   15675: 'Mixinghead 07: Connection 02: Pressure recording: Measuring value outside measuring range', class Mixing Head Warning, trigger "Mixinghead_Pressure_MH7_Con2_DBW320" bit 8
   15676: 'Mixinghead 07: Connection 02: Pressure recording: Warning, value exceeded', class Mixing Head Warning, trigger "Mixinghead_Pressure_MH7_Con2_DBW320" bit 9
   15677: 'Mixinghead 07: Connection 02: Pressure recording: Warning, value undershot', class Mixing Head Warning, trigger "Mixinghead_Pressure_MH7_Con2_DBW320" bit 10
   15678: 'Mixinghead 07: Connection 02: Pressure recording: Fault, value exceeded', class Mixing Head Errors, trigger "Mixinghead_Pressure_MH7_Con2_DBW320" bit 11
   15679: 'Mixinghead 07: Connection 02: Pressure recording: Fault, value undershot', class Mixing Head Errors, trigger "Mixinghead_Pressure_MH7_Con2_DBW320" bit 12
   15680: 'Mixinghead 07: Connection 03: Pressure recording: Measuring value outside measuring range', class Mixing Head Warning, trigger "Mixinghead_Pressure_MH7_Con3_DBW354" bit 8
   15681: 'Mixinghead 07: Connection 03: Pressure recording: Warning, value exceeded', class Mixing Head Warning, trigger "Mixinghead_Pressure_MH7_Con3_DBW354" bit 9
   15682: 'Mixinghead 07: Connection 03: Pressure recording: Warning, value undershot', class Mixing Head Warning, trigger "Mixinghead_Pressure_MH7_Con3_DBW354" bit 10
   15683: 'Mixinghead 07: Connection 03: Pressure recording: Fault, value exceeded', class Mixing Head Errors, trigger "Mixinghead_Pressure_MH7_Con3_DBW354" bit 11
   15684: 'Mixinghead 07: Connection 03: Pressure recording: Fault, value undershot', class Mixing Head Errors, trigger "Mixinghead_Pressure_MH7_Con3_DBW354" bit 12
   15685: 'Mixinghead 07: Connection 04: Pressure recording: Measuring value outside measuring range', class Mixing Head Warning, trigger "Mixinghead_Pressure_MH7_Con4_DBW388" bit 8
   15686: 'Mixinghead 07: Connection 04: Pressure recording: Warning, value exceeded', class Mixing Head Warning, trigger "Mixinghead_Pressure_MH7_Con4_DBW388" bit 9
   15687: 'Mixinghead 07: Connection 04: Pressure recording: Warning, value undershot', class Mixing Head Warning, trigger "Mixinghead_Pressure_MH7_Con4_DBW388" bit 10
   15688: 'Mixinghead 07: Connection 04: Pressure recording: Fault, value exceeded', class Mixing Head Errors, trigger "Mixinghead_Pressure_MH7_Con4_DBW388" bit 11
   15689: 'Mixinghead 07: Connection 04: Pressure recording: Fault, value undershot', class Mixing Head Errors, trigger "Mixinghead_Pressure_MH7_Con4_DBW388" bit 12
   15690: 'Mixinghead 07: Connection 05: Pressure recording: Measuring value outside measuring range', class Mixing Head Warning, trigger "Mixinghead_Pressure_MH7_Con5_DBW422" bit 8
   15691: 'Mixinghead 07: Connection 05: Pressure recording: Warning, value exceeded', class Mixing Head Warning, trigger "Mixinghead_Pressure_MH7_Con5_DBW422" bit 9
   15692: 'Mixinghead 07: Connection 05: Pressure recording: Warning, value undershot', class Mixing Head Warning, trigger "Mixinghead_Pressure_MH7_Con5_DBW422" bit 10
   15693: 'Mixinghead 07: Connection 05: Pressure recording: Fault, value exceeded', class Mixing Head Errors, trigger "Mixinghead_Pressure_MH7_Con5_DBW422" bit 11
   15694: 'Mixinghead 07: Connection 05: Pressure recording: Fault, value undershot', class Mixing Head Errors, trigger "Mixinghead_Pressure_MH7_Con5_DBW422" bit 12
   15695: 'Mixinghead 07: Connection 06: Pressure recording: Measuring value outside measuring range', class Mixing Head Warning, trigger "Mixinghead_Pressure_MH7_Con6_DBW456" bit 8
   15696: 'Mixinghead 07: Connection 06: Pressure recording: Warning, value exceeded', class Mixing Head Warning, trigger "Mixinghead_Pressure_MH7_Con6_DBW456" bit 9
   15697: 'Mixinghead 07: Connection 06: Pressure recording: Warning, value undershot', class Mixing Head Warning, trigger "Mixinghead_Pressure_MH7_Con6_DBW456" bit 10
   15698: 'Mixinghead 07: Connection 06: Pressure recording: Fault, value exceeded', class Mixing Head Errors, trigger "Mixinghead_Pressure_MH7_Con6_DBW456" bit 11
   15699: 'Mixinghead 07: Connection 06: Pressure recording: Fault, value undershot', class Mixing Head Errors, trigger "Mixinghead_Pressure_MH7_Con6_DBW456" bit 12
   15701: 'Mixinghead 08: Mixinghead does not open', class Mixing Head Errors, trigger "Mixinghead_MHControl8_DBW_16" bit 8
   15702: 'Mixinghead 08: Mixinghead does not close', class Mixing Head Errors, trigger "Mixinghead_MHControl8_DBW_16" bit 9
   15703: 'Mixinghead 08: Entry cancelled', class Mixing Head Warning, trigger "Mixinghead_MHControl8_DBW_16" bit 10
   15704: 'Mixinghead 08: Mixinghead open without activation', class Mixing Head Errors, trigger "Mixinghead_MHControl8_DBW_16" bit 11
   15705: 'Mixinghead 08: Mixinghead close during entry', class Mixing Head Warning, trigger "Mixinghead_MHControl8_DBW_16" bit 12
   15706: 'Mixinghead 08: Warning, shot time too short', class Mixing Head Warning, trigger "Mixinghead_MHControl8_DBW_16" bit 13
   15707: 'Mixinghead 08: Warning , shot time too long', class Mixing Head Warning, trigger "Mixinghead_MHControl8_DBW_16" bit 14
   15708: 'Mixinghead 08: Fault, shot time too short', class Mixing Head Warning, trigger "Mixinghead_MHControl8_DBW_16" bit 15
   15709: 'Mixinghead 08: Mixinghead collides when opening or closing', class Mixing Head Warning, trigger "Mixinghead_MHControl8_DBW_16" bit 0
   15710: 'Mixinghead 08: Runtime monitoring when locking mixing head', class Mixing Head Warning, trigger "Mixinghead_MHControl8_DBW_16" bit 1
   15711: 'Mixinghead 08: Runtime monitoring when unlocking mixing head', class Mixing Head Warning, trigger "Mixinghead_MHControl8_DBW_16" bit 2
   15712: 'Mixinghead 08:', class Mixing Head Warning, trigger "Mixinghead_MHControl8_DBW_16" bit 3
   15713: 'Mixinghead 08:', class Mixing Head Warning, trigger "Mixinghead_MHControl8_DBW_16" bit 4
   15714: 'Mixinghead 08:', class Mixing Head Warning, trigger "Mixinghead_MHControl8_DBW_16" bit 5
   15715: 'Mixinghead 08:', class Mixing Head Warning, trigger "Mixinghead_MHControl8_DBW_16" bit 6
   15716: 'Mixinghead 08: Component required in entry is not enabled at this mixing head', class Mixing Head Errors, trigger "Mixinghead_MHControl8_DBW_16" bit 7
   15717: 'Mixinghead 08: Cleaning piston: Moving out too slow', class Mixing Head Errors, trigger "Mixinghead_Cpiston8_DBW_48" bit 8
   15718: 'Mixinghead 08: Cleaning piston: Moving in too slow', class Mixing Head Errors, trigger "Mixinghead_Cpiston8_DBW_48" bit 9
   15719: 'Mixinghead 08: Cleaning piston: Proximity switch defect', class Mixing Head Errors, trigger "Mixinghead_Cpiston8_DBW_48" bit 10
   15720: 'Mixinghead 08: Cleaning piston: Leaves its home position in entry', class Mixing Head Errors, trigger "Mixinghead_Cpiston8_DBW_48" bit 11
   15721: 'Mixinghead 08: Cleaning piston: Not defined', class Mixing Head Warning, trigger "Mixinghead_Cpiston8_DBW_48" bit 12
   15722: 'Mixinghead 08: Cleaning piston:', class Mixing Head Warning, trigger "Mixinghead_Cpiston8_DBW_48" bit 13
   15723: 'Mixinghead 08: Cleaning piston:', class Mixing Head Warning, trigger "Mixinghead_Cpiston8_DBW_48" bit 14
   15724: 'Mixinghead 08: Cleaning piston:', class Mixing Head Warning, trigger "Mixinghead_Cpiston8_DBW_48" bit 15
   15725: 'Mixinghead 08: Cleaning piston: Controller at upper limit', class Mixing Head Warning, trigger "Mixinghead_Cpiston8_DBW_48" bit 0
   15726: 'Mixinghead 08: Cleaning piston: Controller at lower limit', class Mixing Head Warning, trigger "Mixinghead_Cpiston8_DBW_48" bit 1
   15727: 'Mixinghead 08: Cleaning piston:', class Mixing Head Warning, trigger "Mixinghead_Cpiston8_DBW_48" bit 2
   15728: 'Mixinghead 08: Cleaning piston: Front position not reached', class Mixing Head Warning, trigger "Mixinghead_Cpiston8_DBW_48" bit 3
   15729: 'Mixinghead 08: Cleaning piston: Rear position not reached', class Mixing Head Warning, trigger "Mixinghead_Cpiston8_DBW_48" bit 4
   15730: 'Mixinghead 08: Cleaning piston: Home position not reached', class Mixing Head Warning, trigger "Mixinghead_Cpiston8_DBW_48" bit 5
   15731: 'Mixinghead 08: Cleaning piston:', class Mixing Head Warning, trigger "Mixinghead_Cpiston8_DBW_48" bit 6
   15732: 'Mixinghead 08: Cleaning piston:', class Mixing Head Warning, trigger "Mixinghead_Cpiston8_DBW_48" bit 7
   15740: 'Mixinghead 08: Connection 01: Temperature recording: Measuring value outside measuring range', class Mixing Head Warning, trigger "Mixinghead_Temperature_MH8_Con1_DBW84" bit 8
   15741: 'Mixinghead 08: Connection 01: Temperature recording: Warning, value exceeded', class Mixing Head Warning, trigger "Mixinghead_Temperature_MH8_Con1_DBW84" bit 9
   15742: 'Mixinghead 08: Connection 01: Temperature recording: Warning, value undershot', class Mixing Head Warning, trigger "Mixinghead_Temperature_MH8_Con1_DBW84" bit 10
   15743: 'Mixinghead 08: Connection 01: Temperature recording: Fault, value exceeded', class Mixing Head Errors, trigger "Mixinghead_Temperature_MH8_Con1_DBW84" bit 11
   15744: 'Mixinghead 08: Connection 01: Temperature recording: Fault, value undershot', class Mixing Head Errors, trigger "Mixinghead_Temperature_MH8_Con1_DBW84" bit 12
   15745: 'Mixinghead 08: Connection 02: Temperature recording: Measuring value outside measuring range', class Mixing Head Warning, trigger "Mixinghead_Temperature_MH8_Con2_DBW118" bit 8
   15746: 'Mixinghead 08: Connection 02: Temperature recording: Warning, value exceeded', class Mixing Head Warning, trigger "Mixinghead_Temperature_MH8_Con2_DBW118" bit 9
   15747: 'Mixinghead 08: Connection 02: Temperature recording: Warning, value undershot', class Mixing Head Warning, trigger "Mixinghead_Temperature_MH8_Con2_DBW118" bit 10
   15748: 'Mixinghead 08: Connection 02: Temperature recording: Fault, value exceeded', class Mixing Head Errors, trigger "Mixinghead_Temperature_MH8_Con2_DBW118" bit 11
   15749: 'Mixinghead 08: Connection 02: Temperature recording: Fault, value undershot', class Mixing Head Errors, trigger "Mixinghead_Temperature_MH8_Con2_DBW118" bit 12
   15750: 'Mixinghead 08: Connection 03: Temperature recording: Measuring value outside measuring range', class Mixing Head Warning, trigger "Mixinghead_Temperature_MH8_Con3_DBW152" bit 8
   15751: 'Mixinghead 08: Connection 03: Temperature recording: Warning, value exceeded', class Mixing Head Warning, trigger "Mixinghead_Temperature_MH8_Con3_DBW152" bit 9
   15752: 'Mixinghead 08: Connection 03: Temperature recording: Warning, value undershot', class Mixing Head Warning, trigger "Mixinghead_Temperature_MH8_Con3_DBW152" bit 10
   15753: 'Mixinghead 08: Connection 03: Temperature recording: Fault, value exceeded', class Mixing Head Errors, trigger "Mixinghead_Temperature_MH8_Con3_DBW152" bit 11
   15754: 'Mixinghead 08: Connection 03: Temperature recording: Fault, value undershot', class Mixing Head Errors, trigger "Mixinghead_Temperature_MH8_Con3_DBW152" bit 12
   15755: 'Mixinghead 08: Connection 04: Temperature recording: Measuring value outside measuring range', class Mixing Head Warning, trigger "Mixinghead_Temperature_MH8_Con4_DBW186" bit 8
   15756: 'Mixinghead 08: Connection 04: Temperature recording: Warning, value exceeded', class Mixing Head Warning, trigger "Mixinghead_Temperature_MH8_Con4_DBW186" bit 9
   15757: 'Mixinghead 08: Connection 04: Temperature recording: Warning, value undershot', class Mixing Head Warning, trigger "Mixinghead_Temperature_MH8_Con4_DBW186" bit 10
   15758: 'Mixinghead 08: Connection 04: Temperature recording: Fault, value exceeded', class Mixing Head Errors, trigger "Mixinghead_Temperature_MH8_Con4_DBW186" bit 11
   15759: 'Mixinghead 08: Connection 04: Temperature recording: Fault, value undershot', class Mixing Head Errors, trigger "Mixinghead_Temperature_MH8_Con4_DBW186" bit 12
   15760: 'Mixinghead 08: Connection 05: Temperature recording: Measuring value outside measuring range', class Mixing Head Warning, trigger "Mixinghead_Temperature_MH8_Con5_DBW220" bit 8
   15761: 'Mixinghead 08: Connection 05: Temperature recording: Warning, value exceeded', class Mixing Head Warning, trigger "Mixinghead_Temperature_MH8_Con5_DBW220" bit 9
   15762: 'Mixinghead 08: Connection 05: Temperature recording: Warning, value undershot', class Mixing Head Warning, trigger "Mixinghead_Temperature_MH8_Con5_DBW220" bit 10
   15763: 'Mixinghead 08: Connection 05: Temperature recording: Fault, value exceeded', class Mixing Head Errors, trigger "Mixinghead_Temperature_MH8_Con5_DBW220" bit 11
   15764: 'Mixinghead 08: Connection 05: Temperature recording: Fault, value undershot', class Mixing Head Errors, trigger "Mixinghead_Temperature_MH8_Con5_DBW220" bit 12
   15765: 'Mixinghead 08: Connection 06: Temperature recording: Measuring value outside measuring range', class Mixing Head Warning, trigger "Mixinghead_Temperature_MH8_Con6_DBW254" bit 8
   15766: 'Mixinghead 08: Connection 06: Temperature recording: Warning, value exceeded', class Mixing Head Warning, trigger "Mixinghead_Temperature_MH8_Con6_DBW254" bit 9
   15767: 'Mixinghead 08: Connection 06: Temperature recording: Warning, value undershot', class Mixing Head Warning, trigger "Mixinghead_Temperature_MH8_Con6_DBW254" bit 10
   15768: 'Mixinghead 08: Connection 06: Temperature recording: Fault, value exceeded', class Mixing Head Errors, trigger "Mixinghead_Temperature_MH8_Con6_DBW254" bit 11
   15769: 'Mixinghead 08: Connection 06: Temperature recording: Fault, value undershot', class Mixing Head Errors, trigger "Mixinghead_Temperature_MH8_Con6_DBW254" bit 12
   15770: 'Mixinghead 08: Connection 01: Pressure recording: Measuring value outside measuring range', class Mixing Head Warning, trigger "Mixinghead_Pressure_MH8_Con1_DBW288" bit 8
   15771: 'Mixinghead 08: Connection 01: Pressure recording: Warning, value exceeded', class Mixing Head Warning, trigger "Mixinghead_Pressure_MH8_Con1_DBW288" bit 9
   15772: 'Mixinghead 08: Connection 01: Pressure recording: Warning, value undershot', class Mixing Head Warning, trigger "Mixinghead_Pressure_MH8_Con1_DBW288" bit 10
   15773: 'Mixinghead 08: Connection 01: Pressure recording: Fault, value exceeded', class Mixing Head Errors, trigger "Mixinghead_Pressure_MH8_Con1_DBW288" bit 11
   15774: 'Mixinghead 08: Connection 01: Pressure recording: Fault, value undershot', class Mixing Head Errors, trigger "Mixinghead_Pressure_MH8_Con1_DBW288" bit 12
   15775: 'Mixinghead 08: Connection 02: Pressure recording: Measuring value outside measuring range', class Mixing Head Warning, trigger "Mixinghead_Pressure_MH8_Con2_DBW322" bit 8
   15776: 'Mixinghead 08: Connection 02: Pressure recording: Warning, value exceeded', class Mixing Head Warning, trigger "Mixinghead_Pressure_MH8_Con2_DBW322" bit 9
   15777: 'Mixinghead 08: Connection 02: Pressure recording: Warning, value undershot', class Mixing Head Warning, trigger "Mixinghead_Pressure_MH8_Con2_DBW322" bit 10
   15778: 'Mixinghead 08: Connection 02: Pressure recording: Fault, value exceeded', class Mixing Head Errors, trigger "Mixinghead_Pressure_MH8_Con2_DBW322" bit 11
   15779: 'Mixinghead 08: Connection 02: Pressure recording: Fault, value undershot', class Mixing Head Errors, trigger "Mixinghead_Pressure_MH8_Con2_DBW322" bit 12
   15780: 'Mixinghead 08: Connection 03: Pressure recording: Measuring value outside measuring range', class Mixing Head Warning, trigger "Mixinghead_Pressure_MH8_Con3_DBW356" bit 8
   15781: 'Mixinghead 08: Connection 03: Pressure recording: Warning, value exceeded', class Mixing Head Warning, trigger "Mixinghead_Pressure_MH8_Con3_DBW356" bit 9
   15782: 'Mixinghead 08: Connection 03: Pressure recording: Warning, value undershot', class Mixing Head Warning, trigger "Mixinghead_Pressure_MH8_Con3_DBW356" bit 10
   15783: 'Mixinghead 08: Connection 03: Pressure recording: Fault, value exceeded', class Mixing Head Errors, trigger "Mixinghead_Pressure_MH8_Con3_DBW356" bit 11
   15784: 'Mixinghead 08: Connection 03: Pressure recording: Fault, value undershot', class Mixing Head Errors, trigger "Mixinghead_Pressure_MH8_Con3_DBW356" bit 12
   15785: 'Mixinghead 08: Connection 04: Pressure recording: Measuring value outside measuring range', class Mixing Head Warning, trigger "Mixinghead_Pressure_MH8_Con4_DBW390" bit 8
   15786: 'Mixinghead 08: Connection 04: Pressure recording: Warning, value exceeded', class Mixing Head Warning, trigger "Mixinghead_Pressure_MH8_Con4_DBW390" bit 9
   15787: 'Mixinghead 08: Connection 04: Pressure recording: Warning, value undershot', class Mixing Head Warning, trigger "Mixinghead_Pressure_MH8_Con4_DBW390" bit 10
   15788: 'Mixinghead 08: Connection 04: Pressure recording: Fault, value exceeded', class Mixing Head Errors, trigger "Mixinghead_Pressure_MH8_Con4_DBW390" bit 11
   15789: 'Mixinghead 08: Connection 04: Pressure recording: Fault, value undershot', class Mixing Head Errors, trigger "Mixinghead_Pressure_MH8_Con4_DBW390" bit 12
   15790: 'Mixinghead 08: Connection 05: Pressure recording: Measuring value outside measuring range', class Mixing Head Warning, trigger "Mixinghead_Pressure_MH8_Con5_DBW424" bit 8
   15791: 'Mixinghead 08: Connection 05: Pressure recording: Warning, value exceeded', class Mixing Head Warning, trigger "Mixinghead_Pressure_MH8_Con5_DBW424" bit 9
   15792: 'Mixinghead 08: Connection 05: Pressure recording: Warning, value undershot', class Mixing Head Warning, trigger "Mixinghead_Pressure_MH8_Con5_DBW424" bit 10
   15793: 'Mixinghead 08: Connection 05: Pressure recording: Fault, value exceeded', class Mixing Head Errors, trigger "Mixinghead_Pressure_MH8_Con5_DBW424" bit 11
   15794: 'Mixinghead 08: Connection 05: Pressure recording: Fault, value undershot', class Mixing Head Errors, trigger "Mixinghead_Pressure_MH8_Con5_DBW424" bit 12
   15795: 'Mixinghead 08: Connection 06: Pressure recording: Measuring value outside measuring range', class Mixing Head Warning, trigger "Mixinghead_Pressure_MH8_Con6_DBW458" bit 8
   15796: 'Mixinghead 08: Connection 06: Pressure recording: Warning, value exceeded', class Mixing Head Warning, trigger "Mixinghead_Pressure_MH8_Con6_DBW458" bit 9
   15797: 'Mixinghead 08: Connection 06: Pressure recording: Warning, value undershot', class Mixing Head Warning, trigger "Mixinghead_Pressure_MH8_Con6_DBW458" bit 10
   15798: 'Mixinghead 08: Connection 06: Pressure recording: Fault, value exceeded', class Mixing Head Errors, trigger "Mixinghead_Pressure_MH8_Con6_DBW458" bit 11
   15799: 'Mixinghead 08: Connection 06: Pressure recording: Fault, value undershot', class Mixing Head Errors, trigger "Mixinghead_Pressure_MH8_Con6_DBW458" bit 12
   15801: 'Mixinghead 09: Mixinghead does not open', class Mixing Head Errors, trigger "Mixinghead_MHControl9_DBW_18" bit 8
   15802: 'Mixinghead 09: Mixinghead does not close', class Mixing Head Errors, trigger "Mixinghead_MHControl9_DBW_18" bit 9
   15803: 'Mixinghead 09: Entry cancelled', class Mixing Head Warning, trigger "Mixinghead_MHControl9_DBW_18" bit 10
   15804: 'Mixinghead 09: Mixinghead open without activation', class Mixing Head Errors, trigger "Mixinghead_MHControl9_DBW_18" bit 11
   15805: 'Mixinghead 09: Mixinghead close during entry', class Mixing Head Warning, trigger "Mixinghead_MHControl9_DBW_18" bit 12
   15806: 'Mixinghead 09: Warning, shot time too short', class Mixing Head Warning, trigger "Mixinghead_MHControl9_DBW_18" bit 13
   15807: 'Mixinghead 09: Warning , shot time too long', class Mixing Head Warning, trigger "Mixinghead_MHControl9_DBW_18" bit 14
   15808: 'Mixinghead 09: Fault, shot time too short', class Mixing Head Warning, trigger "Mixinghead_MHControl9_DBW_18" bit 15
   15809: 'Mixinghead 09: Mixinghead collides when opening or closing', class Mixing Head Warning, trigger "Mixinghead_MHControl9_DBW_18" bit 0
   15810: 'Mixinghead 09: Runtime monitoring when locking mixing head', class Mixing Head Warning, trigger "Mixinghead_MHControl9_DBW_18" bit 1
   15811: 'Mixinghead 09: Runtime monitoring when unlocking mixing head', class Mixing Head Warning, trigger "Mixinghead_MHControl9_DBW_18" bit 2
   15812: 'Mixinghead 09:', class Mixing Head Warning, trigger "Mixinghead_MHControl9_DBW_18" bit 3
   15813: 'Mixinghead 09:', class Mixing Head Warning, trigger "Mixinghead_MHControl9_DBW_18" bit 4
   15814: 'Mixinghead 09:', class Mixing Head Warning, trigger "Mixinghead_MHControl9_DBW_18" bit 5
   15815: 'Mixinghead 09:', class Mixing Head Warning, trigger "Mixinghead_MHControl9_DBW_18" bit 6
   15816: 'Mixinghead 09: Component required in entry is not enabled at this mixing head', class Mixing Head Errors, trigger "Mixinghead_MHControl9_DBW_18" bit 7
   15817: 'Mixinghead 09: Cleaning piston: Moving out too slow', class Mixing Head Errors, trigger "Mixinghead_Cpiston9_DBW_50" bit 8
   15818: 'Mixinghead 09: Cleaning piston: Moving in too slow', class Mixing Head Errors, trigger "Mixinghead_Cpiston9_DBW_50" bit 9
   15819: 'Mixinghead 09: Cleaning piston: Proximity switch defect', class Mixing Head Errors, trigger "Mixinghead_Cpiston9_DBW_50" bit 10
   15820: 'Mixinghead 09: Cleaning piston: Leaves its home position in entry', class Mixing Head Errors, trigger "Mixinghead_Cpiston9_DBW_50" bit 11
   15821: 'Mixinghead 09: Cleaning piston: Not defined', class Mixing Head Warning, trigger "Mixinghead_Cpiston9_DBW_50" bit 12
   15822: 'Mixinghead 09: Cleaning piston:', class Mixing Head Warning, trigger "Mixinghead_Cpiston9_DBW_50" bit 13
   15823: 'Mixinghead 09: Cleaning piston:', class Mixing Head Warning, trigger "Mixinghead_Cpiston9_DBW_50" bit 14
   15824: 'Mixinghead 09: Cleaning piston:', class Mixing Head Warning, trigger "Mixinghead_Cpiston9_DBW_50" bit 15
   15825: 'Mixinghead 09: Cleaning piston: Controller at upper limit', class Mixing Head Warning, trigger "Mixinghead_Cpiston9_DBW_50" bit 0
   15826: 'Mixinghead 09: Cleaning piston: Controller at lower limit', class Mixing Head Warning, trigger "Mixinghead_Cpiston9_DBW_50" bit 1
   15827: 'Mixinghead 09: Cleaning piston:', class Mixing Head Warning, trigger "Mixinghead_Cpiston9_DBW_50" bit 2
   15828: 'Mixinghead 09: Cleaning piston: Front position not reached', class Mixing Head Warning, trigger "Mixinghead_Cpiston9_DBW_50" bit 3
   15829: 'Mixinghead 09: Cleaning piston: Rear position not reached', class Mixing Head Warning, trigger "Mixinghead_Cpiston9_DBW_50" bit 4
   15830: 'Mixinghead 09: Cleaning piston: Home position not reached', class Mixing Head Warning, trigger "Mixinghead_Cpiston9_DBW_50" bit 5
   15831: 'Mixinghead 09: Cleaning piston:', class Mixing Head Warning, trigger "Mixinghead_Cpiston9_DBW_50" bit 6
   15832: 'Mixinghead 09: Cleaning piston:', class Mixing Head Warning, trigger "Mixinghead_Cpiston9_DBW_50" bit 7
   15840: 'Mixinghead 09: Connection 01: Temperature recording: Measuring value outside measuring range', class Mixing Head Warning, trigger "Mixinghead_Temperature_MH9_Con1_DBW86" bit 8
   15841: 'Mixinghead 09: Connection 01: Temperature recording: Warning, value exceeded', class Mixing Head Warning, trigger "Mixinghead_Temperature_MH9_Con1_DBW86" bit 9
   15842: 'Mixinghead 09: Connection 01: Temperature recording: Warning, value undershot', class Mixing Head Warning, trigger "Mixinghead_Temperature_MH9_Con1_DBW86" bit 10
   15843: 'Mixinghead 09: Connection 01: Temperature recording: Fault, value exceeded', class Mixing Head Errors, trigger "Mixinghead_Temperature_MH9_Con1_DBW86" bit 11
   15844: 'Mixinghead 09: Connection 01: Temperature recording: Fault, value undershot', class Mixing Head Errors, trigger "Mixinghead_Temperature_MH9_Con1_DBW86" bit 12
   15845: 'Mixinghead 09: Connection 02: Temperature recording: Measuring value outside measuring range', class Mixing Head Warning, trigger "Mixinghead_Temperature_MH9_Con2_DBW120" bit 8
   15846: 'Mixinghead 09: Connection 02: Temperature recording: Warning, value exceeded', class Mixing Head Warning, trigger "Mixinghead_Temperature_MH9_Con2_DBW120" bit 9
   15847: 'Mixinghead 09: Connection 02: Temperature recording: Warning, value undershot', class Mixing Head Warning, trigger "Mixinghead_Temperature_MH9_Con2_DBW120" bit 10
   15848: 'Mixinghead 09: Connection 02: Temperature recording: Fault, value exceeded', class Mixing Head Errors, trigger "Mixinghead_Temperature_MH9_Con2_DBW120" bit 11
   15849: 'Mixinghead 09: Connection 02: Temperature recording: Fault, value undershot', class Mixing Head Errors, trigger "Mixinghead_Temperature_MH9_Con2_DBW120" bit 12
   15850: 'Mixinghead 09: Connection 03: Temperature recording: Measuring value outside measuring range', class Mixing Head Warning, trigger "Mixinghead_Temperature_MH9_Con3_DBW154" bit 8
   15851: 'Mixinghead 09: Connection 03: Temperature recording: Warning, value exceeded', class Mixing Head Warning, trigger "Mixinghead_Temperature_MH9_Con3_DBW154" bit 9
   15852: 'Mixinghead 09: Connection 03: Temperature recording: Warning, value undershot', class Mixing Head Warning, trigger "Mixinghead_Temperature_MH9_Con3_DBW154" bit 10
   15853: 'Mixinghead 09: Connection 03: Temperature recording: Fault, value exceeded', class Mixing Head Errors, trigger "Mixinghead_Temperature_MH9_Con3_DBW154" bit 11
   15854: 'Mixinghead 09: Connection 03: Temperature recording: Fault, value undershot', class Mixing Head Errors, trigger "Mixinghead_Temperature_MH9_Con3_DBW154" bit 12
   15855: 'Mixinghead 09: Connection 04: Temperature recording: Measuring value outside measuring range', class Mixing Head Warning, trigger "Mixinghead_Temperature_MH9_Con4_DBW188" bit 8
   15856: 'Mixinghead 09: Connection 04: Temperature recording: Warning, value exceeded', class Mixing Head Warning, trigger "Mixinghead_Temperature_MH9_Con4_DBW188" bit 9
   15857: 'Mixinghead 09: Connection 04: Temperature recording: Warning, value undershot', class Mixing Head Warning, trigger "Mixinghead_Temperature_MH9_Con4_DBW188" bit 10
   15858: 'Mixinghead 09: Connection 04: Temperature recording: Fault, value exceeded', class Mixing Head Errors, trigger "Mixinghead_Temperature_MH9_Con4_DBW188" bit 11
   15859: 'Mixinghead 09: Connection 04: Temperature recording: Fault, value undershot', class Mixing Head Errors, trigger "Mixinghead_Temperature_MH9_Con4_DBW188" bit 12
   15860: 'Mixinghead 09: Connection 05: Temperature recording: Measuring value outside measuring range', class Mixing Head Warning, trigger "Mixinghead_Temperature_MH9_Con5_DBW222" bit 8
   15861: 'Mixinghead 09: Connection 05: Temperature recording: Warning, value exceeded', class Mixing Head Warning, trigger "Mixinghead_Temperature_MH9_Con5_DBW222" bit 9
   15862: 'Mixinghead 09: Connection 05: Temperature recording: Warning, value undershot', class Mixing Head Warning, trigger "Mixinghead_Temperature_MH9_Con5_DBW222" bit 10
   15863: 'Mixinghead 09: Connection 05: Temperature recording: Fault, value exceeded', class Mixing Head Errors, trigger "Mixinghead_Temperature_MH9_Con5_DBW222" bit 11
   15864: 'Mixinghead 09: Connection 05: Temperature recording: Fault, value undershot', class Mixing Head Errors, trigger "Mixinghead_Temperature_MH9_Con5_DBW222" bit 12
   15865: 'Mixinghead 09: Connection 06: Temperature recording: Measuring value outside measuring range', class Mixing Head Warning, trigger "Mixinghead_Temperature_MH9_Con6_DBW256" bit 8
   15866: 'Mixinghead 09: Connection 06: Temperature recording: Warning, value exceeded', class Mixing Head Warning, trigger "Mixinghead_Temperature_MH9_Con6_DBW256" bit 9
   15867: 'Mixinghead 09: Connection 06: Temperature recording: Warning, value undershot', class Mixing Head Warning, trigger "Mixinghead_Temperature_MH9_Con6_DBW256" bit 10
   15868: 'Mixinghead 09: Connection 06: Temperature recording: Fault, value exceeded', class Mixing Head Errors, trigger "Mixinghead_Temperature_MH9_Con6_DBW256" bit 11
   15869: 'Mixinghead 09: Connection 06: Temperature recording: Fault, value undershot', class Mixing Head Errors, trigger "Mixinghead_Temperature_MH9_Con6_DBW256" bit 12
   15870: 'Mixinghead 09: Connection 01: Pressure recording: Measuring value outside measuring range', class Mixing Head Warning, trigger "Mixinghead_Pressure_MH9_Con1_DBW290" bit 8
   15871: 'Mixinghead 09: Connection 01: Pressure recording: Warning, value exceeded', class Mixing Head Warning, trigger "Mixinghead_Pressure_MH9_Con1_DBW290" bit 9
   15872: 'Mixinghead 09: Connection 01: Pressure recording: Warning, value undershot', class Mixing Head Warning, trigger "Mixinghead_Pressure_MH9_Con1_DBW290" bit 10
   15873: 'Mixinghead 09: Connection 01: Pressure recording: Fault, value exceeded', class Mixing Head Errors, trigger "Mixinghead_Pressure_MH9_Con1_DBW290" bit 11
   15874: 'Mixinghead 09: Connection 01: Pressure recording: Fault, value undershot', class Mixing Head Errors, trigger "Mixinghead_Pressure_MH9_Con1_DBW290" bit 12
   15875: 'Mixinghead 09: Connection 02: Pressure recording: Measuring value outside measuring range', class Mixing Head Warning, trigger "Mixinghead_Pressure_MH9_Con2_DBW324" bit 8
   15876: 'Mixinghead 09: Connection 02: Pressure recording: Warning, value exceeded', class Mixing Head Warning, trigger "Mixinghead_Pressure_MH9_Con2_DBW324" bit 9
   15877: 'Mixinghead 09: Connection 02: Pressure recording: Warning, value undershot', class Mixing Head Warning, trigger "Mixinghead_Pressure_MH9_Con2_DBW324" bit 10
   15878: 'Mixinghead 09: Connection 02: Pressure recording: Fault, value exceeded', class Mixing Head Errors, trigger "Mixinghead_Pressure_MH9_Con2_DBW324" bit 11
   15879: 'Mixinghead 09: Connection 02: Pressure recording: Fault, value undershot', class Mixing Head Errors, trigger "Mixinghead_Pressure_MH9_Con2_DBW324" bit 12
   15880: 'Mixinghead 09: Connection 03: Pressure recording: Measuring value outside measuring range', class Mixing Head Warning, trigger "Mixinghead_Pressure_MH9_Con3_DBW358" bit 8
   15881: 'Mixinghead 09: Connection 03: Pressure recording: Warning, value exceeded', class Mixing Head Warning, trigger "Mixinghead_Pressure_MH9_Con3_DBW358" bit 9
   15882: 'Mixinghead 09: Connection 03: Pressure recording: Warning, value undershot', class Mixing Head Warning, trigger "Mixinghead_Pressure_MH9_Con3_DBW358" bit 10
   15883: 'Mixinghead 09: Connection 03: Pressure recording: Fault, value exceeded', class Mixing Head Errors, trigger "Mixinghead_Pressure_MH9_Con3_DBW358" bit 11
   15884: 'Mixinghead 09: Connection 03: Pressure recording: Fault, value undershot', class Mixing Head Errors, trigger "Mixinghead_Pressure_MH9_Con3_DBW358" bit 12
   15885: 'Mixinghead 09: Connection 04: Pressure recording: Measuring value outside measuring range', class Mixing Head Warning, trigger "Mixinghead_Pressure_MH9_Con4_DBW392" bit 8
   15886: 'Mixinghead 09: Connection 04: Pressure recording: Warning, value exceeded', class Mixing Head Warning, trigger "Mixinghead_Pressure_MH9_Con4_DBW392" bit 9
   15887: 'Mixinghead 09: Connection 04: Pressure recording: Warning, value undershot', class Mixing Head Warning, trigger "Mixinghead_Pressure_MH9_Con4_DBW392" bit 10
   15888: 'Mixinghead 09: Connection 04: Pressure recording: Fault, value exceeded', class Mixing Head Errors, trigger "Mixinghead_Pressure_MH9_Con4_DBW392" bit 11
   15889: 'Mixinghead 09: Connection 04: Pressure recording: Fault, value undershot', class Mixing Head Errors, trigger "Mixinghead_Pressure_MH9_Con4_DBW392" bit 12
   15890: 'Mixinghead 09: Connection 05: Pressure recording: Measuring value outside measuring range', class Mixing Head Warning, trigger "Mixinghead_Pressure_MH9_Con5_DBW426" bit 8
   15891: 'Mixinghead 09: Connection 05: Pressure recording: Warning, value exceeded', class Mixing Head Warning, trigger "Mixinghead_Pressure_MH9_Con5_DBW426" bit 9
   15892: 'Mixinghead 09: Connection 05: Pressure recording: Warning, value undershot', class Mixing Head Warning, trigger "Mixinghead_Pressure_MH9_Con5_DBW426" bit 10
   15893: 'Mixinghead 09: Connection 05: Pressure recording: Fault, value exceeded', class Mixing Head Errors, trigger "Mixinghead_Pressure_MH9_Con5_DBW426" bit 11
   15894: 'Mixinghead 09: Connection 05: Pressure recording: Fault, value undershot', class Mixing Head Errors, trigger "Mixinghead_Pressure_MH9_Con5_DBW426" bit 12
   15895: 'Mixinghead 09: Connection 06: Pressure recording: Measuring value outside measuring range', class Mixing Head Warning, trigger "Mixinghead_Pressure_MH9_Con6_DBW460" bit 0
   15896: 'Mixinghead 09: Connection 06: Pressure recording: Warning, value exceeded', class Mixing Head Warning, trigger "Mixinghead_Pressure_MH9_Con6_DBW460" bit 1
   15897: 'Mixinghead 09: Connection 06: Pressure recording: Warning, value undershot', class Mixing Head Warning, trigger "Mixinghead_Pressure_MH9_Con6_DBW460" bit 2
   15898: 'Mixinghead 09: Connection 06: Pressure recording: Fault, value exceeded', class Mixing Head Errors, trigger "Mixinghead_Pressure_MH9_Con6_DBW460" bit 3
   15899: 'Mixinghead 09: Connection 06: Pressure recording: Fault, value undershot', class Mixing Head Errors, trigger "Mixinghead_Pressure_MH9_Con6_DBW460" bit 4
   15901: 'Mixinghead 10: Mixinghead does not open', class Mixing Head Errors, trigger "Mixinghead_MHControl10_DBW_20" bit 8
   15902: 'Mixinghead 10: Mixinghead does not close', class Mixing Head Errors, trigger "Mixinghead_MHControl10_DBW_20" bit 9
   15903: 'Mixinghead 10: Entry cancelled', class Mixing Head Warning, trigger "Mixinghead_MHControl10_DBW_20" bit 10
   15904: 'Mixinghead 10: Mixinghead open without activation', class Mixing Head Errors, trigger "Mixinghead_MHControl10_DBW_20" bit 11
   15905: 'Mixinghead 10: Mixinghead close during entry', class Mixing Head Warning, trigger "Mixinghead_MHControl10_DBW_20" bit 12
   15906: 'Mixinghead 10: Warning, shot time too short', class Mixing Head Warning, trigger "Mixinghead_MHControl10_DBW_20" bit 13
   15907: 'Mixinghead 10: Warning , shot time too long', class Mixing Head Warning, trigger "Mixinghead_MHControl10_DBW_20" bit 14
   15908: 'Mixinghead 10: Fault, shot time too short', class Mixing Head Warning, trigger "Mixinghead_MHControl10_DBW_20" bit 15
   15909: 'Mixinghead 10: Mixinghead collides when opening or closing', class Mixing Head Warning, trigger "Mixinghead_MHControl10_DBW_20" bit 0
   15910: 'Mixinghead 10: Runtime monitoring when locking mixing head', class Mixing Head Warning, trigger "Mixinghead_MHControl10_DBW_20" bit 1
   15911: 'Mixinghead 10: Runtime monitoring when unlocking mixing head', class Mixing Head Warning, trigger "Mixinghead_MHControl10_DBW_20" bit 2
   15912: 'Mixinghead 10:', class Mixing Head Warning, trigger "Mixinghead_MHControl10_DBW_20" bit 3
   15913: 'Mixinghead 10:', class Mixing Head Warning, trigger "Mixinghead_MHControl10_DBW_20" bit 4
   15914: 'Mixinghead 10:', class Mixing Head Warning, trigger "Mixinghead_MHControl10_DBW_20" bit 5
   15915: 'Mixinghead 10:', class Mixing Head Warning, trigger "Mixinghead_MHControl10_DBW_20" bit 6
   15916: 'Mixinghead 10: Component required in entry is not enabled at this mixing head', class Mixing Head Errors, trigger "Mixinghead_MHControl10_DBW_20" bit 7
   15917: 'Mixinghead 10: Cleaning piston: Moving out too slow', class Mixing Head Errors, trigger "Mixinghead_Cpiston10_DBW_52" bit 8
   15918: 'Mixinghead 10: Cleaning piston: Moving in too slow', class Mixing Head Errors, trigger "Mixinghead_Cpiston10_DBW_52" bit 9
   15919: 'Mixinghead 10: Cleaning piston: Proximity switch defect', class Mixing Head Errors, trigger "Mixinghead_Cpiston10_DBW_52" bit 10
   15920: 'Mixinghead 10: Cleaning piston: Leaves its home position in entry', class Mixing Head Errors, trigger "Mixinghead_Cpiston10_DBW_52" bit 11
   15921: 'Mixinghead 10: Cleaning piston: Not defined', class Mixing Head Warning, trigger "Mixinghead_Cpiston10_DBW_52" bit 12
   15922: 'Mixinghead 10: Cleaning piston:', class Mixing Head Warning, trigger "Mixinghead_Cpiston10_DBW_52" bit 13
   15923: 'Mixinghead 10: Cleaning piston:', class Mixing Head Warning, trigger "Mixinghead_Cpiston10_DBW_52" bit 14
   15924: 'Mixinghead 10: Cleaning piston:', class Mixing Head Warning, trigger "Mixinghead_Cpiston10_DBW_52" bit 15
   15925: 'Mixinghead 10: Cleaning piston: Controller at upper limit', class Mixing Head Warning, trigger "Mixinghead_Cpiston10_DBW_52" bit 0
   15926: 'Mixinghead 10: Cleaning piston: Controller at lower limit', class Mixing Head Warning, trigger "Mixinghead_Cpiston10_DBW_52" bit 1
   15927: 'Mixinghead 10: Cleaning piston:', class Mixing Head Warning, trigger "Mixinghead_Cpiston10_DBW_52" bit 2
   15928: 'Mixinghead 10: Cleaning piston: Front position not reached', class Mixing Head Warning, trigger "Mixinghead_Cpiston10_DBW_52" bit 3
   15929: 'Mixinghead 10: Cleaning piston: Rear position not reached', class Mixing Head Warning, trigger "Mixinghead_Cpiston10_DBW_52" bit 4
   15930: 'Mixinghead 10: Cleaning piston: Home position not reached', class Mixing Head Warning, trigger "Mixinghead_Cpiston10_DBW_52" bit 5
   15931: 'Mixinghead 10: Cleaning piston:', class Mixing Head Warning, trigger "Mixinghead_Cpiston10_DBW_52" bit 6
   15932: 'Mixinghead 10: Cleaning piston:', class Mixing Head Warning, trigger "Mixinghead_Cpiston10_DBW_52" bit 7
   15940: 'Mixinghead 10: Connection 01: Temperature recording: Measuring value outside measuring range', class Mixing Head Warning, trigger "Mixinghead_Temperature_MH10_Con1_DBW88" bit 8
   15941: 'Mixinghead 10: Connection 01: Temperature recording: Warning, value exceeded', class Mixing Head Warning, trigger "Mixinghead_Temperature_MH10_Con1_DBW88" bit 9
   15942: 'Mixinghead 10: Connection 01: Temperature recording: Warning, value undershot', class Mixing Head Warning, trigger "Mixinghead_Temperature_MH10_Con1_DBW88" bit 10
   15943: 'Mixinghead 10: Connection 01: Temperature recording: Fault, value exceeded', class Mixing Head Errors, trigger "Mixinghead_Temperature_MH10_Con1_DBW88" bit 11
   15944: 'Mixinghead 10: Connection 01: Temperature recording: Fault, value undershot', class Mixing Head Errors, trigger "Mixinghead_Temperature_MH10_Con1_DBW88" bit 12
   15945: 'Mixinghead 10: Connection 02: Temperature recording: Measuring value outside measuring range', class Mixing Head Warning, trigger "Mixinghead_Temperature_MH10_Con2_DBW122" bit 8
   15946: 'Mixinghead 10: Connection 02: Temperature recording: Warning, value exceeded', class Mixing Head Warning, trigger "Mixinghead_Temperature_MH10_Con2_DBW122" bit 9
   15947: 'Mixinghead 10: Connection 02: Temperature recording: Warning, value undershot', class Mixing Head Warning, trigger "Mixinghead_Temperature_MH10_Con2_DBW122" bit 10
   15948: 'Mixinghead 10: Connection 02: Temperature recording: Fault, value exceeded', class Mixing Head Errors, trigger "Mixinghead_Temperature_MH10_Con2_DBW122" bit 11
   15949: 'Mixinghead 10: Connection 02: Temperature recording: Fault, value undershot', class Mixing Head Errors, trigger "Mixinghead_Temperature_MH10_Con2_DBW122" bit 12
   15950: 'Mixinghead 10: Connection 03: Temperature recording: Measuring value outside measuring range', class Mixing Head Warning, trigger "Mixinghead_Temperature_MH10_Con3_DBW156" bit 8
   15951: 'Mixinghead 10: Connection 03: Temperature recording: Warning, value exceeded', class Mixing Head Warning, trigger "Mixinghead_Temperature_MH10_Con3_DBW156" bit 9
   15952: 'Mixinghead 10: Connection 03: Temperature recording: Warning, value undershot', class Mixing Head Warning, trigger "Mixinghead_Temperature_MH10_Con3_DBW156" bit 10
   15953: 'Mixinghead 10: Connection 03: Temperature recording: Fault, value exceeded', class Mixing Head Errors, trigger "Mixinghead_Temperature_MH10_Con3_DBW156" bit 11
   15954: 'Mixinghead 10: Connection 03: Temperature recording: Fault, value undershot', class Mixing Head Errors, trigger "Mixinghead_Temperature_MH10_Con3_DBW156" bit 12
   15955: 'Mixinghead 10: Connection 04: Temperature recording: Measuring value outside measuring range', class Mixing Head Warning, trigger "Mixinghead_Temperature_MH10_Con4_DBW190" bit 8
   15956: 'Mixinghead 10: Connection 04: Temperature recording: Warning, value exceeded', class Mixing Head Warning, trigger "Mixinghead_Temperature_MH10_Con4_DBW190" bit 9
   15957: 'Mixinghead 10: Connection 04: Temperature recording: Warning, value undershot', class Mixing Head Warning, trigger "Mixinghead_Temperature_MH10_Con4_DBW190" bit 10
   15958: 'Mixinghead 10: Connection 04: Temperature recording: Fault, value exceeded', class Mixing Head Errors, trigger "Mixinghead_Temperature_MH10_Con4_DBW190" bit 11
   15959: 'Mixinghead 10: Connection 04: Temperature recording: Fault, value undershot', class Mixing Head Errors, trigger "Mixinghead_Temperature_MH10_Con4_DBW190" bit 12
   15960: 'Mixinghead 10: Connection 05: Temperature recording: Measuring value outside measuring range', class Mixing Head Warning, trigger "Mixinghead_Temperature_MH10_Con5_DBW224" bit 8
   15961: 'Mixinghead 10: Connection 05: Temperature recording: Warning, value exceeded', class Mixing Head Warning, trigger "Mixinghead_Temperature_MH10_Con5_DBW224" bit 9
   15962: 'Mixinghead 10: Connection 05: Temperature recording: Warning, value undershot', class Mixing Head Warning, trigger "Mixinghead_Temperature_MH10_Con5_DBW224" bit 10
   15963: 'Mixinghead 10: Connection 05: Temperature recording: Fault, value exceeded', class Mixing Head Errors, trigger "Mixinghead_Temperature_MH10_Con5_DBW224" bit 11
   15964: 'Mixinghead 10: Connection 05: Temperature recording: Fault, value undershot', class Mixing Head Errors, trigger "Mixinghead_Temperature_MH10_Con5_DBW224" bit 12
   15965: 'Mixinghead 10: Connection 06: Temperature recording: Measuring value outside measuring range', class Mixing Head Warning, trigger "Mixinghead_Temperature_MH10_Con6_DBW258" bit 8
   15966: 'Mixinghead 10: Connection 06: Temperature recording: Warning, value exceeded', class Mixing Head Warning, trigger "Mixinghead_Temperature_MH10_Con6_DBW258" bit 9
   15967: 'Mixinghead 10: Connection 06: Temperature recording: Warning, value undershot', class Mixing Head Warning, trigger "Mixinghead_Temperature_MH10_Con6_DBW258" bit 10
   15968: 'Mixinghead 10: Connection 06: Temperature recording: Fault, value exceeded', class Mixing Head Errors, trigger "Mixinghead_Temperature_MH10_Con6_DBW258" bit 11
   15969: 'Mixinghead 10: Connection 06: Temperature recording: Fault, value undershot', class Mixing Head Errors, trigger "Mixinghead_Temperature_MH10_Con6_DBW258" bit 12
   15970: 'Mixinghead 10: Connection 01: Pressure recording: Measuring value outside measuring range', class Mixing Head Warning, trigger "Mixinghead_Pressure_MH10_Con1_DBW292" bit 8
   15971: 'Mixinghead 10: Connection 01: Pressure recording: Warning, value exceeded', class Mixing Head Warning, trigger "Mixinghead_Pressure_MH10_Con1_DBW292" bit 9
   15972: 'Mixinghead 10: Connection 01: Pressure recording: Warning, value undershot', class Mixing Head Warning, trigger "Mixinghead_Pressure_MH10_Con1_DBW292" bit 10
   15973: 'Mixinghead 10: Connection 01: Pressure recording: Fault, value exceeded', class Mixing Head Errors, trigger "Mixinghead_Pressure_MH10_Con1_DBW292" bit 11
   15974: 'Mixinghead 10: Connection 01: Pressure recording: Fault, value undershot', class Mixing Head Errors, trigger "Mixinghead_Pressure_MH10_Con1_DBW292" bit 12
   15975: 'Mixinghead 10: Connection 02: Pressure recording: Measuring value outside measuring range', class Mixing Head Warning, trigger "Mixinghead_Pressure_MH10_Con2_DBW326" bit 8
   15976: 'Mixinghead 10: Connection 02: Pressure recording: Warning, value exceeded', class Mixing Head Warning, trigger "Mixinghead_Pressure_MH10_Con2_DBW326" bit 9
   15977: 'Mixinghead 10: Connection 02: Pressure recording: Warning, value undershot', class Mixing Head Warning, trigger "Mixinghead_Pressure_MH10_Con2_DBW326" bit 10
   15978: 'Mixinghead 10: Connection 02: Pressure recording: Fault, value exceeded', class Mixing Head Errors, trigger "Mixinghead_Pressure_MH10_Con2_DBW326" bit 11
   15979: 'Mixinghead 10: Connection 02: Pressure recording: Fault, value undershot', class Mixing Head Errors, trigger "Mixinghead_Pressure_MH10_Con2_DBW326" bit 12
   15980: 'Mixinghead 10: Connection 03: Pressure recording: Measuring value outside measuring range', class Mixing Head Warning, trigger "Mixinghead_Pressure_MH10_Con3_DBW360" bit 8
   15981: 'Mixinghead 10: Connection 03: Pressure recording: Warning, value exceeded', class Mixing Head Warning, trigger "Mixinghead_Pressure_MH10_Con3_DBW360" bit 9
   15982: 'Mixinghead 10: Connection 03: Pressure recording: Warning, value undershot', class Mixing Head Warning, trigger "Mixinghead_Pressure_MH10_Con3_DBW360" bit 10
   15983: 'Mixinghead 10: Connection 03: Pressure recording: Fault, value exceeded', class Mixing Head Errors, trigger "Mixinghead_Pressure_MH10_Con3_DBW360" bit 11